   "Carrier_42_G120DControlWord.4" AT %I2460.4 : Bool;   // Bit_04_EN_RAMP
   "Carrier_42_G120DControlWord.5" AT %I2460.5 : Bool;   // Bit_05_START_RAMP
   "Carrier_42_G120DControlWord.6" AT %I2460.6 : Bool;   // Bit_06_SETPOINT
   "Carrier_42_G120DControlWord.7" AT %I2460.7 : Bool;   // Bit_07_RESET
   "Carrier_42_G120DControlWord.8" AT %I2461.0 : Bool;   // Bit_08_JOG_R
   "Carrier_42_G120DControlWord.9" AT %I2461.1 : Bool;   // Bit_09_JOG_L
   "Carrier_42_G120DControlWord.10" AT %I2461.2 : Bool;   // Bit_10_CONTR_PLC
   "Carrier_42_G120DControlWord.11" AT %I2461.3 : Bool;   // Bit_11_REVERSE
   "Carrier_42_G120DControlWord.12" AT %I2461.4 : Bool;   // Bit_12_BRAKE_RELEASE
   "Carrier_42_G120DControlWord.13" AT %I2461.5 : Bool;   // Bit_13_DDS
   "Carrier_42_G120DControlWord.14" AT %I2461.6 : Bool;   // Bit_14_DO0
   "Carrier_42_G120DControlWord.15" AT %I2461.7 : Bool;   // Bit_15_DO1
   "Carrier_42_G120DStatusWord" AT %IW2462 : Word;   // G120D_ZSW1_STATUS
   "Carrier_42_G120DStatusWord.0" AT %I2462.0 : Bool;   // Bit_00_READY_RUN
   "Carrier_42_G120DStatusWord.1" AT %I2462.1 : Bool;   // Bit_01_READY_ON
   "Carrier_42_G120DStatusWord.2" AT %I2462.2 : Bool;   // Bit_02_ENABLE
   "Carrier_42_G120DStatusWord.3" AT %I2462.3 : Bool;   // Bit_03_FAULT
   "Carrier_42_G120DStatusWord.4" AT %I2462.4 : Bool;   // Bit_04_OFF2
   "Carrier_42_G120DStatusWord.5" AT %I2462.5 : Bool;   // Bit_05_OFF3
   "Carrier_42_G120DStatusWord.6" AT %I2462.6 : Bool;   // Bit_06_LOCK_OUT
   "Carrier_42_G120DStatusWord.7" AT %I2462.7 : Bool;   // Bit_07_WARN
   "Carrier_42_G120DStatusWord.8" AT %I2463.0 : Bool;   // Bit_08_NO_DEVIATION
   "Carrier_42_G120DStatusWord.9" AT %I2463.1 : Bool;   // Bit_09_CONTR_PLC
   "Carrier_42_G120DStatusWord.10" AT %I2463.2 : Bool;   // Bit_10_F_MAX
   "Carrier_42_G120DStatusWord.11" AT %I2463.3 : Bool;   // Bit_11_LIMIT_REACHED
   "Carrier_42_G120DStatusWord.12" AT %I2463.4 : Bool;   // Bit_12_BRAKE_OPEN
   "Carrier_42_G120DStatusWord.13" AT %I2463.5 : Bool;   // Bit_13_NO_OVERTEMP
   "Carrier_42_G120DStatusWord.14" AT %I2463.6 : Bool;   // Bit_14_CW_CCW
   "Carrier_42_G120DStatusWord.15" AT %I2463.7 : Bool;   // Bit_15_OVERL
   "Carrier_42_Slot2_Input" AT %IW2464 : Word;   // SLOT 2 INPUT WORD
   "Carrier_42_CrashDetectSW" AT %I2464.0 : Bool;   // CRASH DETECT SW
   "Carrier_42_SpareSafetyInput(2_1)" AT %I2464.1 : Bool;   // SPARE SAFETY INPUT
   "Carrier_42_SpareSafetyInput(2_2)" AT %I2464.2 : Bool;   // SPARE SAFETY INPUT
   "Carrier_42_SpareSafetyInput(2_3)" AT %I2464.3 : Bool;   // SPARE SAFETY INPUT
   "Carrier_42_SpareSafetyInput(2_4)" AT %I2464.4 : Bool;   // SPARE SAFETY INPUT
   "Carrier_42_SpareSafetyInput(2_5)" AT %I2464.5 : Bool;   // SPARE SAFETY INPUT
   "Carrier_42_SpareSafetyInput(2_6)" AT %I2464.6 : Bool;   // SPARE SAFETY INPUT
   "Carrier_42_SpareSafetyInput(2_7)" AT %I2464.7 : Bool;   // SPARE SAFETY INPUT
   "Carrier_42_Slot3_SafetyOutput" AT %IW2465 : Word;   // SLOT 3 SAFETY OUTPUT WORD
   "Carrier_42_Crash_Detect_OK" AT %I2465.0 : Bool;   // CARRIER CRASH DETECT
   "Carrier_42_SpareSafetyOutput(3_1)" AT %I2465.1 : Bool;   // SPARE SAFETY OUTPUT
   "Carrier_42_SpareSafetyOutput(3_2)" AT %I2465.2 : Bool;   // SPARE SAFETY OUTPUT
   "Carrier_42_SpareSafetyOutput(3_3)" AT %I2465.3 : Bool;   // SPARE SAFETY OUTPUT
   "Carrier_42_SpareSafetyOutput(3_4)" AT %I2465.4 : Bool;   // SPARE SAFETY OUTPUT
   "Carrier_42_SpareSafetyOutput(3_5)" AT %I2465.5 : Bool;   // SPARE SAFETY OUTPUT
   "Carrier_42_SpareSafetyOutput(3_6)" AT %I2465.6 : Bool;   // SPARE SAFETY OUTPUT
   "Carrier_42_SpareSafetyOutput(3_7)" AT %I2465.7 : Bool;   // SPARE SAFETY OUTPUT
   "Carrier_42_Slot4_Input" AT %IW2466 : Word;   // SLOT 4 INPUT WORD
   "Carrier_42_480VPowerOn_MDCB1" AT %I2466.0 : Bool;   // 480 VAC POWER ON MDCB 1
   "Carrier_42_SpareInput(4_1)" AT %I2466.1 : Bool;   // SPARE INPUT
   "Carrier_42_SpareInput(4_2)" AT %I2466.2 : Bool;   // SPARE INPUT
   "Carrier_42_SitopSelectStatus" AT %I2466.3 : Bool;   // SITOP SELECT STATUS
   "Carrier_42_DCsupplyOnPSCB2" AT %I2466.4 : Bool;   // DC SUPPLY ON PSCB 2
   "Carrier_42_SpareInput(4_5)" AT %I2466.5 : Bool;   // SPARE INPUT
   "Carrier_42_SpareInput(4_6)" AT %I2466.6 : Bool;   // SPARE INPUT
   "Carrier_42_SpareInput(4_7)" AT %I2466.7 : Bool;   // SPARE INPUT
   "Carrier_42_PB1_ProdHoldLH" AT %I2467.0 : Bool;   // PB 1 PRODUCTION HOLD LH
   "Carrier_42_PB2_ResetLH" AT %I2467.1 : Bool;   // PB 2 RESET LH
   "Carrier_42_PB3_ProdHoldRH" AT %I2467.2 : Bool;   // PB 3 PRODUCTION HOLD RH
   "Carrier_42_PB4_ResetRH" AT %I2467.3 : Bool;   // PB 4 RESET RH
   "Carrier_42_SpareInput(4_14)" AT %I2467.4 : Bool;   // SPARE INPUT
   "Carrier_42_SpareInput(4_15)" AT %I2467.5 : Bool;   // SPARE INPUT
   "Carrier_42_SpareInput(4_16)" AT %I2467.6 : Bool;   // SPARE INPUT
   "Carrier_42_SpareInput(4_17)" AT %I2467.7 : Bool;   // SPARE INPUT
   "Carrier_42_Slot5_Output" AT %IW2468 : Word;   // SLOT 5 OUTPUT WORD
   "Carrier_42_IRD400_HMI_24VDC_ENABLE" AT %I2468.0 : Bool;   // IRD 400 PANEL HMI 24V DC POWER
   "Carrier_42_FaultLight_LH" AT %I2468.1 : Bool;   // FAULT LIGHT LH
   "Carrier_42_RunLight_LH" AT %I2468.2 : Bool;   // RUN LIGHT LH
   "Carrier_42_FaultLight_RH" AT %I2468.3 : Bool;   // FAULT LIGHT RH
   "Carrier_42_RunLight_RH" AT %I2468.4 : Bool;   // RUN LIGHT RH
   "Carrier_42_SpareOutput(5_5)" AT %I2468.5 : Bool;   // SPARE OUTPUT
   "Carrier_42_SpareOutput(5_6)" AT %I2468.6 : Bool;   // SPARE OUTPUT
   "Carrier_42_SpareOutput(5_7)" AT %I2468.7 : Bool;   // SPARE OUTPUT
   "Carrier_42_ActualSpeed" AT %IW2470 : Word;   // ACTUAL SPEED
   "Carrier_42_CarrierDriveAlarm" AT %IW2472 : Word;   // CARRIER DRIVE ALARM
   "Carrier_42_CarrierDriveWarning" AT %IW2474 : Word;   // CARRIER DRIVE WARNING
   "Carrier_43_Status" AT %IW2500 : Word;   // CARRIER STATUS WORD
   "Carrier_43_Status.0" AT %I2500.0 : Bool;   // HEARTBEAT
   "Carrier_43_Status.1" AT %I2500.1 : Bool;   // MANUAL
   "Carrier_43_Status.2" AT %I2500.2 : Bool;   // IN_AUTO
   "Carrier_43_Status.3" AT %I2500.3 : Bool;   // POSITIONING_COMPLETE
   "Carrier_43_Status.4" AT %I2500.4 : Bool;   // PRODUCTION HOLD
   "Carrier_43_Status.5" AT %I2500.5 : Bool;   // CARRIER MOVING FORWARD
   "Carrier_43_Status.6" AT %I2500.6 : Bool;   // CARRIER MOVING REVERSE
   "Carrier_43_Status.7" AT %I2500.7 : Bool;   // CARRIER FAULT
   "Carrier_43_Status.8" AT %I2501.0 : Bool;   // CRASH DETECT TRIPPED
   "Carrier_43_Status.9" AT %I2501.1 : Bool;
   "Carrier_43_Status.10" AT %I2501.2 : Bool;
   "Carrier_43_Status.11" AT %I2501.3 : Bool;
   "Carrier_43_Status.12" AT %I2501.4 : Bool;
   "Carrier_43_Status.13" AT %I2501.5 : Bool;
   "Carrier_43_Status.14" AT %I2501.6 : Bool;
   "Carrier_43_Status.15" AT %I2501.7 : Bool;
   "Carrier_43_SDCFaultCode" AT %IW2502 : Word;   // SDC FAULT CODE
   "Carrier_43_CarrierPosition" AT %ID2504 : DWord;   // CARRIER POSITION
   "Carrier_43_CarrierNumber" AT %IW2508 : Word;   // CARRIER NUMBER
   "Carrier_43_G120DControlWord" AT %IW2510 : Word;   // G120D_STW1_CONTROL
   "Carrier_43_G120DControlWord.0" AT %I2510.0 : Bool;   // Bit_00_ON
   "Carrier_43_G120DControlWord.1" AT %I2510.1 : Bool;   // Bit_01_AUS2_INH
   "Carrier_43_G120DControlWord.2" AT %I2510.2 : Bool;   // Bit_02_AUS3_STOP
   "Carrier_43_G120DControlWord.3" AT %I2510.3 : Bool;   // Bit_03_EN
   "Carrier_43_G120DControlWord.4" AT %I2510.4 : Bool;   // Bit_04_EN_RAMP
   "Carrier_43_G120DControlWord.5" AT %I2510.5 : Bool;   // Bit_05_START_RAMP
   "Carrier_43_G120DControlWord.6" AT %I2510.6 : Bool;   // Bit_06_SETPOINT
   "Carrier_43_G120DControlWord.7" AT %I2510.7 : Bool;   // Bit_07_RESET
   "Carrier_43_G120DControlWord.8" AT %I2511.0 : Bool;   // Bit_08_JOG_R
   "Carrier_43_G120DControlWord.9" AT %I2511.1 : Bool;   // Bit_09_JOG_L
   "Carrier_43_G120DControlWord.10" AT %I2511.2 : Bool;   // Bit_10_CONTR_PLC
   "Carrier_43_G120DControlWord.11" AT %I2511.3 : Bool;   // Bit_11_REVERSE
   "Carrier_43_G120DControlWord.12" AT %I2511.4 : Bool;   // Bit_12_BRAKE_RELEASE
   "Carrier_43_G120DControlWord.13" AT %I2511.5 : Bool;   // Bit_13_DDS
   "Carrier_43_G120DControlWord.14" AT %I2511.6 : Bool;   // Bit_14_DO0
   "Carrier_43_G120DControlWord.15" AT %I2511.7 : Bool;   // Bit_15_DO1
   "Carrier_43_G120DStatusWord" AT %IW2512 : Word;   // G120D_ZSW1_STATUS
   "Carrier_43_G120DStatusWord.0" AT %I2512.0 : Bool;   // Bit_00_READY_RUN
   "Carrier_43_G120DStatusWord.1" AT %I2512.1 : Bool;   // Bit_01_READY_ON
   "Carrier_43_G120DStatusWord.2" AT %I2512.2 : Bool;   // Bit_02_ENABLE
   "Carrier_43_G120DStatusWord.3" AT %I2512.3 : Bool;   // Bit_03_FAULT
   "Carrier_43_G120DStatusWord.4" AT %I2512.4 : Bool;   // Bit_04_OFF2
   "Carrier_43_G120DStatusWord.5" AT %I2512.5 : Bool;   // Bit_05_OFF3
   "Carrier_43_G120DStatusWord.6" AT %I2512.6 : Bool;   // Bit_06_LOCK_OUT
   "Carrier_43_G120DStatusWord.7" AT %I2512.7 : Bool;   // Bit_07_WARN
   "Carrier_43_G120DStatusWord.8" AT %I2513.0 : Bool;   // Bit_08_NO_DEVIATION
   "Carrier_43_G120DStatusWord.9" AT %I2513.1 : Bool;   // Bit_09_CONTR_PLC
   "Carrier_43_G120DStatusWord.10" AT %I2513.2 : Bool;   // Bit_10_F_MAX
   "Carrier_43_G120DStatusWord.11" AT %I2513.3 : Bool;   // Bit_11_LIMIT_REACHED
   "Carrier_43_G120DStatusWord.12" AT %I2513.4 : Bool;   // Bit_12_BRAKE_OPEN
   "Carrier_43_G120DStatusWord.13" AT %I2513.5 : Bool;   // Bit_13_NO_OVERTEMP
   "Carrier_43_G120DStatusWord.14" AT %I2513.6 : Bool;   // Bit_14_CW_CCW
   "Carrier_43_G120DStatusWord.15" AT %I2513.7 : Bool;   // Bit_15_OVERL
   "Carrier_43_Slot2_Input" AT %IW2514 : Word;   // SLOT 2 INPUT WORD
   "Carrier_43_CrashDetectSW" AT %I2514.0 : Bool;   // CRASH DETECT SW
   "Carrier_43_SpareSafetyInput(2_1)" AT %I2514.1 : Bool;   // SPARE SAFETY INPUT
   "Carrier_43_SpareSafetyInput(2_2)" AT %I2514.2 : Bool;   // SPARE SAFETY INPUT
   "Carrier_43_SpareSafetyInput(2_3)" AT %I2514.3 : Bool;   // SPARE SAFETY INPUT
   "Carrier_43_SpareSafetyInput(2_4)" AT %I2514.4 : Bool;   // SPARE SAFETY INPUT
   "Carrier_43_SpareSafetyInput(2_5)" AT %I2514.5 : Bool;   // SPARE SAFETY INPUT
   "Carrier_43_SpareSafetyInput(2_6)" AT %I2514.6 : Bool;   // SPARE SAFETY INPUT
   "Carrier_43_SpareSafetyInput(2_7)" AT %I2514.7 : Bool;   // SPARE SAFETY INPUT
   "Carrier_43_Slot3_SafetyOutput" AT %IW2515 : Word;   // SLOT 3 SAFETY OUTPUT WORD
   "Carrier_43_Crash_Detect_OK" AT %I2515.0 : Bool;   // CARRIER CRASH DETECT
   "Carrier_43_SpareSafetyOutput(3_1)" AT %I2515.1 : Bool;   // SPARE SAFETY OUTPUT
   "Carrier_43_SpareSafetyOutput(3_2)" AT %I2515.2 : Bool;   // SPARE SAFETY OUTPUT
   "Carrier_43_SpareSafetyOutput(3_3)" AT %I2515.3 : Bool;   // SPARE SAFETY OUTPUT
   "Carrier_43_SpareSafetyOutput(3_4)" AT %I2515.4 : Bool;   // SPARE SAFETY OUTPUT
   "Carrier_43_SpareSafetyOutput(3_5)" AT %I2515.5 : Bool;   // SPARE SAFETY OUTPUT
   "Carrier_43_SpareSafetyOutput(3_6)" AT %I2515.6 : Bool;   // SPARE SAFETY OUTPUT
   "Carrier_43_SpareSafetyOutput(3_7)" AT %I2515.7 : Bool;   // SPARE SAFETY OUTPUT
   "Carrier_43_Slot4_Input" AT %IW2516 : Word;   // SLOT 4 INPUT WORD
   "Carrier_43_480VPowerOn_MDCB1" AT %I2516.0 : Bool;   // 480 VAC POWER ON MDCB 1
   "Carrier_43_SpareInput(4_1)" AT %I2516.1 : Bool;   // SPARE INPUT
   "Carrier_43_SpareInput(4_2)" AT %I2516.2 : Bool;   // SPARE INPUT
   "Carrier_43_SitopSelectStatus" AT %I2516.3 : Bool;   // SITOP SELECT STATUS
   "Carrier_43_DCsupplyOnPSCB2" AT %I2516.4 : Bool;   // DC SUPPLY ON PSCB 2
   "Carrier_43_SpareInput(4_5)" AT %I2516.5 : Bool;   // SPARE INPUT
   "Carrier_43_SpareInput(4_6)" AT %I2516.6 : Bool;   // SPARE INPUT
   "Carrier_43_SpareInput(4_7)" AT %I2516.7 : Bool;   // SPARE INPUT
   "Carrier_43_PB1_ProdHoldLH" AT %I2517.0 : Bool;   // PB 1 PRODUCTION HOLD LH
   "Carrier_43_PB2_ResetLH" AT %I2517.1 : Bool;   // PB 2 RESET LH
   "Carrier_43_PB3_ProdHoldRH" AT %I2517.2 : Bool;   // PB 3 PRODUCTION HOLD RH
   "Carrier_43_PB4_ResetRH" AT %I2517.3 : Bool;   // PB 4 RESET RH
   "Carrier_43_SpareInput(4_14)" AT %I2517.4 : Bool;   // SPARE INPUT
   "Carrier_43_SpareInput(4_15)" AT %I2517.5 : Bool;   // SPARE INPUT
   "Carrier_43_SpareInput(4_16)" AT %I2517.6 : Bool;   // SPARE INPUT
   "Carrier_43_SpareInput(4_17)" AT %I2517.7 : Bool;   // SPARE INPUT
   "Carrier_43_Slot5_Output" AT %IW2518 : Word;   // SLOT 5 OUTPUT WORD
   "Carrier_43_IRD400_HMI_24VDC_ENABLE" AT %I2518.0 : Bool;   // IRD 400 PANEL HMI 24V DC POWER
   "Carrier_43_FaultLight_LH" AT %I2518.1 : Bool;   // FAULT LIGHT LH
   "Carrier_43_RunLight_LH" AT %I2518.2 : Bool;   // RUN LIGHT LH
   "Carrier_43_FaultLight_RH" AT %I2518.3 : Bool;   // FAULT LIGHT RH
   "Carrier_43_RunLight_RH" AT %I2518.4 : Bool;   // RUN LIGHT RH
   "Carrier_43_SpareOutput(5_5)" AT %I2518.5 : Bool;   // SPARE OUTPUT
   "Carrier_43_SpareOutput(5_6)" AT %I2518.6 : Bool;   // SPARE OUTPUT
   "Carrier_43_SpareOutput(5_7)" AT %I2518.7 : Bool;   // SPARE OUTPUT
   "Carrier_43_ActualSpeed" AT %IW2520 : Word;   // ACTUAL SPEED
   "Carrier_43_CarrierDriveAlarm" AT %IW2522 : Word;   // CARRIER DRIVE ALARM
   "Carrier_43_CarrierDriveWarning" AT %IW2524 : Word;   // CARRIER DRIVE WARNING
   "Carrier_44_Status" AT %IW2550 : Word;   // CARRIER STATUS WORD
   "Carrier_44_Status.0" AT %I2550.0 : Bool;   // HEARTBEAT
   "Carrier_44_Status.1" AT %I2550.1 : Bool;   // MANUAL
   "Carrier_44_Status.2" AT %I2550.2 : Bool;   // IN_AUTO
   "Carrier_44_Status.3" AT %I2550.3 : Bool;   // POSITIONING_COMPLETE
   "Carrier_44_Status.4" AT %I2550.4 : Bool;   // PRODUCTION HOLD
   "Carrier_44_Status.5" AT %I2550.5 : Bool;   // CARRIER MOVING FORWARD
   "Carrier_44_Status.6" AT %I2550.6 : Bool;   // CARRIER MOVING REVERSE
   "Carrier_44_Status.7" AT %I2550.7 : Bool;   // CARRIER FAULT
   "Carrier_44_Status.8" AT %I2551.0 : Bool;   // CRASH DETECT TRIPPED
   "Carrier_44_Status.9" AT %I2551.1 : Bool;
   "Carrier_44_Status.10" AT %I2551.2 : Bool;
   "Carrier_44_Status.11" AT %I2551.3 : Bool;
   "Carrier_44_Status.12" AT %I2551.4 : Bool;
   "Carrier_44_Status.13" AT %I2551.5 : Bool;
   "Carrier_44_Status.14" AT %I2551.6 : Bool;
   "Carrier_44_Status.15" AT %I2551.7 : Bool;
   "Carrier_44_SDCFaultCode" AT %IW2552 : Word;   // SDC FAULT CODE
   "Carrier_44_CarrierPosition" AT %ID2554 : DWord;   // CARRIER POSITION
   "Carrier_44_CarrierNumber" AT %IW2558 : Word;   // CARRIER NUMBER
   "Carrier_44_G120DControlWord" AT %IW2560 : Word;   // G120D_STW1_CONTROL
   "Carrier_44_G120DControlWord.0" AT %I2560.0 : Bool;   // Bit_00_ON
   "Carrier_44_G120DControlWord.1" AT %I2560.1 : Bool;   // Bit_01_AUS2_INH
   "Carrier_44_G120DControlWord.2" AT %I2560.2 : Bool;   // Bit_02_AUS3_STOP
   "Carrier_44_G120DControlWord.3" AT %I2560.3 : Bool;   // Bit_03_EN
   "Carrier_44_G120DControlWord.4" AT %I2560.4 : Bool;   // Bit_04_EN_RAMP
   "Carrier_44_G120DControlWord.5" AT %I2560.5 : Bool;   // Bit_05_START_RAMP
   "Carrier_44_G120DControlWord.6" AT %I2560.6 : Bool;   // Bit_06_SETPOINT
   "Carrier_44_G120DControlWord.7" AT %I2560.7 : Bool;   // Bit_07_RESET
   "Carrier_44_G120DControlWord.8" AT %I2561.0 : Bool;   // Bit_08_JOG_R
   "Carrier_44_G120DControlWord.9" AT %I2561.1 : Bool;   // Bit_09_JOG_L
   "Carrier_44_G120DControlWord.10" AT %I2561.2 : Bool;   // Bit_10_CONTR_PLC
   "Carrier_44_G120DControlWord.11" AT %I2561.3 : Bool;   // Bit_11_REVERSE
   "Carrier_44_G120DControlWord.12" AT %I2561.4 : Bool;   // Bit_12_BRAKE_RELEASE
   "Carrier_44_G120DControlWord.13" AT %I2561.5 : Bool;   // Bit_13_DDS
   "Carrier_44_G120DControlWord.14" AT %I2561.6 : Bool;   // Bit_14_DO0
   "Carrier_44_G120DControlWord.15" AT %I2561.7 : Bool;   // Bit_15_DO1
   "Carrier_44_G120DStatusWord" AT %IW2562 : Word;   // G120D_ZSW1_STATUS
   "Carrier_44_G120DStatusWord.0" AT %I2562.0 : Bool;   // Bit_00_READY_RUN
   "Carrier_44_G120DStatusWord.1" AT %I2562.1 : Bool;   // Bit_01_READY_ON
   "Carrier_44_G120DStatusWord.2" AT %I2562.2 : Bool;   // Bit_02_ENABLE
   "Carrier_44_G120DStatusWord.3" AT %I2562.3 : Bool;   // Bit_03_FAULT
   "Carrier_44_G120DStatusWord.4" AT %I2562.4 : Bool;   // Bit_04_OFF2
   "Carrier_44_G120DStatusWord.5" AT %I2562.5 : Bool;   // Bit_05_OFF3
   "Carrier_44_G120DStatusWord.6" AT %I2562.6 : Bool;   // Bit_06_LOCK_OUT
   "Carrier_44_G120DStatusWord.7" AT %I2562.7 : Bool;   // Bit_07_WARN
   "Carrier_44_G120DStatusWord.8" AT %I2563.0 : Bool;   // Bit_08_NO_DEVIATION
   "Carrier_44_G120DStatusWord.9" AT %I2563.1 : Bool;   // Bit_09_CONTR_PLC
   "Carrier_44_G120DStatusWord.10" AT %I2563.2 : Bool;   // Bit_10_F_MAX
   "Carrier_44_G120DStatusWord.11" AT %I2563.3 : Bool;   // Bit_11_LIMIT_REACHED
   "Carrier_44_G120DStatusWord.12" AT %I2563.4 : Bool;   // Bit_12_BRAKE_OPEN
   "Carrier_44_G120DStatusWord.13" AT %I2563.5 : Bool;   // Bit_13_NO_OVERTEMP
   "Carrier_44_G120DStatusWord.14" AT %I2563.6 : Bool;   // Bit_14_CW_CCW
   "Carrier_44_G120DStatusWord.15" AT %I2563.7 : Bool;   // Bit_15_OVERL
   "Carrier_44_Slot2_Input" AT %IW2564 : Word;   // SLOT 2 INPUT WORD
   "Carrier_44_CrashDetectSW" AT %I2564.0 : Bool;   // CRASH DETECT SW
   "Carrier_44_SpareSafetyInput(2_1)" AT %I2564.1 : Bool;   // SPARE SAFETY INPUT
   "Carrier_44_SpareSafetyInput(2_2)" AT %I2564.2 : Bool;   // SPARE SAFETY INPUT
   "Carrier_44_SpareSafetyInput(2_3)" AT %I2564.3 : Bool;   // SPARE SAFETY INPUT
   "Carrier_44_SpareSafetyInput(2_4)" AT %I2564.4 : Bool;   // SPARE SAFETY INPUT
   "Carrier_44_SpareSafetyInput(2_5)" AT %I2564.5 : Bool;   // SPARE SAFETY INPUT
   "Carrier_44_SpareSafetyInput(2_6)" AT %I2564.6 : Bool;   // SPARE SAFETY INPUT
   "Carrier_44_SpareSafetyInput(2_7)" AT %I2564.7 : Bool;   // SPARE SAFETY INPUT
   "Carrier_44_Slot3_SafetyOutput" AT %IW2565 : Word;   // SLOT 3 SAFETY OUTPUT WORD
   "Carrier_44_Crash_Detect_OK" AT %I2565.0 : Bool;   // CARRIER CRASH DETECT
   "Carrier_44_SpareSafetyOutput(3_1)" AT %I2565.1 : Bool;   // SPARE SAFETY OUTPUT
   "Carrier_44_SpareSafetyOutput(3_2)" AT %I2565.2 : Bool;   // SPARE SAFETY OUTPUT
   "Carrier_44_SpareSafetyOutput(3_3)" AT %I2565.3 : Bool;   // SPARE SAFETY OUTPUT
   "Carrier_44_SpareSafetyOutput(3_4)" AT %I2565.4 : Bool;   // SPARE SAFETY OUTPUT
   "Carrier_44_SpareSafetyOutput(3_5)" AT %I2565.5 : Bool;   // SPARE SAFETY OUTPUT
   "Carrier_44_SpareSafetyOutput(3_6)" AT %I2565.6 : Bool;   // SPARE SAFETY OUTPUT
   "Carrier_44_SpareSafetyOutput(3_7)" AT %I2565.7 : Bool;   // SPARE SAFETY OUTPUT
   "Carrier_44_Slot4_Input" AT %IW2566 : Word;   // SLOT 4 INPUT WORD
   "Carrier_44_480VPowerOn_MDCB1" AT %I2566.0 : Bool;   // 480 VAC POWER ON MDCB 1
   "Carrier_44_SpareInput(4_1)" AT %I2566.1 : Bool;   // SPARE INPUT
   "Carrier_44_SpareInput(4_2)" AT %I2566.2 : Bool;   // SPARE INPUT
   "Carrier_44_SitopSelectStatus" AT %I2566.3 : Bool;   // SITOP SELECT STATUS
   "Carrier_44_DCsupplyOnPSCB2" AT %I2566.4 : Bool;   // DC SUPPLY ON PSCB 2
   "Carrier_44_SpareInput(4_5)" AT %I2566.5 : Bool;   // SPARE INPUT
   "Carrier_44_SpareInput(4_6)" AT %I2566.6 : Bool;   // SPARE INPUT
   "Carrier_44_SpareInput(4_7)" AT %I2566.7 : Bool;   // SPARE INPUT
   "Carrier_44_PB1_ProdHoldLH" AT %I2567.0 : Bool;   // PB 1 PRODUCTION HOLD LH
   "Carrier_44_PB2_ResetLH" AT %I2567.1 : Bool;   // PB 2 RESET LH
   "Carrier_44_PB3_ProdHoldRH" AT %I2567.2 : Bool;   // PB 3 PRODUCTION HOLD RH
   "Carrier_44_PB4_ResetRH" AT %I2567.3 : Bool;   // PB 4 RESET RH
   "Carrier_44_SpareInput(4_14)" AT %I2567.4 : Bool;   // SPARE INPUT
   "Carrier_44_SpareInput(4_15)" AT %I2567.5 : Bool;   // SPARE INPUT
   "Carrier_44_SpareInput(4_16)" AT %I2567.6 : Bool;   // SPARE INPUT
   "Carrier_44_SpareInput(4_17)" AT %I2567.7 : Bool;   // SPARE INPUT
   "Carrier_44_Slot5_Output" AT %IW2568 : Word;   // SLOT 5 OUTPUT WORD
   "Carrier_44_IRD400_HMI_24VDC_ENABLE" AT %I2568.0 : Bool;   // IRD 400 PANEL HMI 24V DC POWER
   "Carrier_44_FaultLight_LH" AT %I2568.1 : Bool;   // FAULT LIGHT LH
   "Carrier_44_RunLight_LH" AT %I2568.2 : Bool;   // RUN LIGHT LH
   "Carrier_44_FaultLight_RH" AT %I2568.3 : Bool;   // FAULT LIGHT RH
   "Carrier_44_RunLight_RH" AT %I2568.4 : Bool;   // RUN LIGHT RH
   "Carrier_44_SpareOutput(5_5)" AT %I2568.5 : Bool;   // SPARE OUTPUT
   "Carrier_44_SpareOutput(5_6)" AT %I2568.6 : Bool;   // SPARE OUTPUT
   "Carrier_44_SpareOutput(5_7)" AT %I2568.7 : Bool;   // SPARE OUTPUT
   "Carrier_44_ActualSpeed" AT %IW2570 : Word;   // ACTUAL SPEED
   "Carrier_44_CarrierDriveAlarm" AT %IW2572 : Word;   // CARRIER DRIVE ALARM
   "Carrier_44_CarrierDriveWarning" AT %IW2574 : Word;   // CARRIER DRIVE WARNING
   "Carrier_45_Status" AT %IW2600 : Word;   // CARRIER STATUS WORD
   "Carrier_45_Status.0" AT %I2600.0 : Bool;   // HEARTBEAT
   "Carrier_45_Status.1" AT %I2600.1 : Bool;   // MANUAL
   "Carrier_45_Status.2" AT %I2600.2 : Bool;   // IN_AUTO
   "Carrier_45_Status.3" AT %I2600.3 : Bool;   // POSITIONING_COMPLETE
   "Carrier_45_Status.4" AT %I2600.4 : Bool;   // PRODUCTION HOLD
   "Carrier_45_Status.5" AT %I2600.5 : Bool;   // CARRIER MOVING FORWARD
   "Carrier_45_Status.6" AT %I2600.6 : Bool;   // CARRIER MOVING REVERSE
   "Carrier_45_Status.7" AT %I2600.7 : Bool;   // CARRIER FAULT
   "Carrier_45_Status.8" AT %I2601.0 : Bool;   // CRASH DETECT TRIPPED
   "Carrier_45_Status.9" AT %I2601.1 : Bool;
   "Carrier_45_Status.10" AT %I2601.2 : Bool;
   "Carrier_45_Status.11" AT %I2601.3 : Bool;
   "Carrier_45_Status.12" AT %I2601.4 : Bool;
   "Carrier_45_Status.13" AT %I2601.5 : Bool;
   "Carrier_45_Status.14" AT %I2601.6 : Bool;
   "Carrier_45_Status.15" AT %I2601.7 : Bool;
   "Carrier_45_SDCFaultCode" AT %IW2602 : Word;   // SDC FAULT CODE
   "Carrier_45_CarrierPosition" AT %ID2604 : DWord;   // CARRIER POSITION
   "Carrier_45_CarrierNumber" AT %IW2608 : Word;   // CARRIER NUMBER
   "Carrier_45_G120DControlWord" AT %IW2610 : Word;   // G120D_STW1_CONTROL
   "Carrier_45_G120DControlWord.0" AT %I2610.0 : Bool;   // Bit_00_ON
   "Carrier_45_G120DControlWord.1" AT %I2610.1 : Bool;   // Bit_01_AUS2_INH
   "Carrier_45_G120DControlWord.2" AT %I2610.2 : Bool;   // Bit_02_AUS3_STOP
   "Carrier_45_G120DControlWord.3" AT %I2610.3 : Bool;   // Bit_03_EN
   "Carrier_45_G120DControlWord.4" AT %I2610.4 : Bool;   // Bit_04_EN_RAMP
   "Carrier_45_G120DControlWord.5" AT %I2610.5 : Bool;   // Bit_05_START_RAMP
   "Carrier_45_G120DControlWord.6" AT %I2610.6 : Bool;   // Bit_06_SETPOINT
   "Carrier_45_G120DControlWord.7" AT %I2610.7 : Bool;   // Bit_07_RESET
   "Carrier_45_G120DControlWord.8" AT %I2611.0 : Bool;   // Bit_08_JOG_R
   "Carrier_45_G120DControlWord.9" AT %I2611.1 : Bool;   // Bit_09_JOG_L
   "Carrier_45_G120DControlWord.10" AT %I2611.2 : Bool;   // Bit_10_CONTR_PLC
   "Carrier_45_G120DControlWord.11" AT %I2611.3 : Bool;   // Bit_11_REVERSE
   "Carrier_45_G120DControlWord.12" AT %I2611.4 : Bool;   // Bit_12_BRAKE_RELEASE
   "Carrier_45_G120DControlWord.13" AT %I2611.5 : Bool;   // Bit_13_DDS
   "Carrier_45_G120DControlWord.14" AT %I2611.6 : Bool;   // Bit_14_DO0
   "Carrier_45_G120DControlWord.15" AT %I2611.7 : Bool;   // Bit_15_DO1
   "Carrier_45_G120DStatusWord" AT %IW2612 : Word;   // G120D_ZSW1_STATUS
   "Carrier_45_G120DStatusWord.0" AT %I2612.0 : Bool;   // Bit_00_READY_RUN
   "Carrier_45_G120DStatusWord.1" AT %I2612.1 : Bool;   // Bit_01_READY_ON
   "Carrier_45_G120DStatusWord.2" AT %I2612.2 : Bool;   // Bit_02_ENABLE
   "Carrier_45_G120DStatusWord.3" AT %I2612.3 : Bool;   // Bit_03_FAULT
   "Carrier_45_G120DStatusWord.4" AT %I2612.4 : Bool;   // Bit_04_OFF2
   "Carrier_45_G120DStatusWord.5" AT %I2612.5 : Bool;   // Bit_05_OFF3
   "Carrier_45_G120DStatusWord.6" AT %I2612.6 : Bool;   // Bit_06_LOCK_OUT
   "Carrier_45_G120DStatusWord.7" AT %I2612.7 : Bool;   // Bit_07_WARN
   "Carrier_45_G120DStatusWord.8" AT %I2613.0 : Bool;   // Bit_08_NO_DEVIATION
   "Carrier_45_G120DStatusWord.9" AT %I2613.1 : Bool;   // Bit_09_CONTR_PLC
   "Carrier_45_G120DStatusWord.10" AT %I2613.2 : Bool;   // Bit_10_F_MAX
   "Carrier_45_G120DStatusWord.11" AT %I2613.3 : Bool;   // Bit_11_LIMIT_REACHED
   "Carrier_45_G120DStatusWord.12" AT %I2613.4 : Bool;   // Bit_12_BRAKE_OPEN
   "Carrier_45_G120DStatusWord.13" AT %I2613.5 : Bool;   // Bit_13_NO_OVERTEMP
   "Carrier_45_G120DStatusWord.14" AT %I2613.6 : Bool;   // Bit_14_CW_CCW
   "Carrier_45_G120DStatusWord.15" AT %I2613.7 : Bool;   // Bit_15_OVERL
   "Carrier_45_Slot2_Input" AT %IW2614 : Word;   // SLOT 2 INPUT WORD
   "Carrier_45_CrashDetectSW" AT %I2614.0 : Bool;   // CRASH DETECT SW
   "Carrier_45_SpareSafetyInput(2_1)" AT %I2614.1 : Bool;   // SPARE SAFETY INPUT
   "Carrier_45_SpareSafetyInput(2_2)" AT %I2614.2 : Bool;   // SPARE SAFETY INPUT
   "Carrier_45_SpareSafetyInput(2_3)" AT %I2614.3 : Bool;   // SPARE SAFETY INPUT
   "Carrier_45_SpareSafetyInput(2_4)" AT %I2614.4 : Bool;   // SPARE SAFETY INPUT
   "Carrier_45_SpareSafetyInput(2_5)" AT %I2614.5 : Bool;   // SPARE SAFETY INPUT
   "Carrier_45_SpareSafetyInput(2_6)" AT %I2614.6 : Bool;   // SPARE SAFETY INPUT
   "Carrier_45_SpareSafetyInput(2_7)" AT %I2614.7 : Bool;   // SPARE SAFETY INPUT
   "Carrier_45_Slot3_SafetyOutput" AT %IW2615 : Word;   // SLOT 3 SAFETY OUTPUT WORD
   "Carrier_45_Crash_Detect_OK" AT %I2615.0 : Bool;   // CARRIER CRASH DETECT
   "Carrier_45_SpareSafetyOutput(3_1)" AT %I2615.1 : Bool;   // SPARE SAFETY OUTPUT
   "Carrier_45_SpareSafetyOutput(3_2)" AT %I2615.2 : Bool;   // SPARE SAFETY OUTPUT
   "Carrier_45_SpareSafetyOutput(3_3)" AT %I2615.3 : Bool;   // SPARE SAFETY OUTPUT
   "Carrier_45_SpareSafetyOutput(3_4)" AT %I2615.4 : Bool;   // SPARE SAFETY OUTPUT
   "Carrier_45_SpareSafetyOutput(3_5)" AT %I2615.5 : Bool;   // SPARE SAFETY OUTPUT
   "Carrier_45_SpareSafetyOutput(3_6)" AT %I2615.6 : Bool;   // SPARE SAFETY OUTPUT
   "Carrier_45_SpareSafetyOutput(3_7)" AT %I2615.7 : Bool;   // SPARE SAFETY OUTPUT
   "Carrier_45_Slot4_Input" AT %IW2616 : Word;   // SLOT 4 INPUT WORD
   "Carrier_45_480VPowerOn_MDCB1" AT %I2616.0 : Bool;   // 480 VAC POWER ON MDCB 1
   "Carrier_45_SpareInput(4_1)" AT %I2616.1 : Bool;   // SPARE INPUT
   "Carrier_45_SpareInput(4_2)" AT %I2616.2 : Bool;   // SPARE INPUT
   "Carrier_45_SitopSelectStatus" AT %I2616.3 : Bool;   // SITOP SELECT STATUS
   "Carrier_45_DCsupplyOnPSCB2" AT %I2616.4 : Bool;   // DC SUPPLY ON PSCB 2
   "Carrier_45_SpareInput(4_5)" AT %I2616.5 : Bool;   // SPARE INPUT
   "Carrier_45_SpareInput(4_6)" AT %I2616.6 : Bool;   // SPARE INPUT
   "Carrier_45_SpareInput(4_7)" AT %I2616.7 : Bool;   // SPARE INPUT
   "Carrier_45_PB1_ProdHoldLH" AT %I2617.0 : Bool;   // PB 1 PRODUCTION HOLD LH
   "Carrier_45_PB2_ResetLH" AT %I2617.1 : Bool;   // PB 2 RESET LH
   "Carrier_45_PB3_ProdHoldRH" AT %I2617.2 : Bool;   // PB 3 PRODUCTION HOLD RH
   "Carrier_45_PB4_ResetRH" AT %I2617.3 : Bool;   // PB 4 RESET RH
   "Carrier_45_SpareInput(4_14)" AT %I2617.4 : Bool;   // SPARE INPUT
   "Carrier_45_SpareInput(4_15)" AT %I2617.5 : Bool;   // SPARE INPUT
   "Carrier_45_SpareInput(4_16)" AT %I2617.6 : Bool;   // SPARE INPUT
   "Carrier_45_SpareInput(4_17)" AT %I2617.7 : Bool;   // SPARE INPUT
   "Carrier_45_Slot5_Output" AT %IW2618 : Word;   // SLOT 5 OUTPUT WORD
   "Carrier_45_IRD400_HMI_24VDC_ENABLE" AT %I2618.0 : Bool;   // IRD 400 PANEL HMI 24V DC POWER
   "Carrier_45_FaultLight_LH" AT %I2618.1 : Bool;   // FAULT LIGHT LH
   "Carrier_45_RunLight_LH" AT %I2618.2 : Bool;   // RUN LIGHT LH
   "Carrier_45_FaultLight_RH" AT %I2618.3 : Bool;   // FAULT LIGHT RH
   "Carrier_45_RunLight_RH" AT %I2618.4 : Bool;   // RUN LIGHT RH
   "Carrier_45_SpareOutput(5_5)" AT %I2618.5 : Bool;   // SPARE OUTPUT
   "Carrier_45_SpareOutput(5_6)" AT %I2618.6 : Bool;   // SPARE OUTPUT
   "Carrier_45_SpareOutput(5_7)" AT %I2618.7 : Bool;   // SPARE OUTPUT
   "Carrier_45_ActualSpeed" AT %IW2620 : Word;   // ACTUAL SPEED
   "Carrier_45_CarrierDriveAlarm" AT %IW2622 : Word;   // CARRIER DRIVE ALARM
   "Carrier_45_CarrierDriveWarning" AT %IW2624 : Word;   // CARRIER DRIVE WARNING
   "Carrier_46_Status" AT %IW2650 : Word;   // CARRIER STATUS WORD
   "Carrier_46_Status.0" AT %I2650.0 : Bool;   // HEARTBEAT
   "Carrier_46_Status.1" AT %I2650.1 : Bool;   // MANUAL
   "Carrier_46_Status.2" AT %I2650.2 : Bool;   // IN_AUTO
   "Carrier_46_Status.3" AT %I2650.3 : Bool;   // POSITIONING_COMPLETE
   "Carrier_46_Status.4" AT %I2650.4 : Bool;   // PRODUCTION HOLD
   "Carrier_46_Status.5" AT %I2650.5 : Bool;   // CARRIER MOVING FORWARD
   "Carrier_46_Status.6" AT %I2650.6 : Bool;   // CARRIER MOVING REVERSE
   "Carrier_46_Status.7" AT %I2650.7 : Bool;   // CARRIER FAULT
   "Carrier_46_Status.8" AT %I2651.0 : Bool;   // CRASH DETECT TRIPPED
   "Carrier_46_Status.9" AT %I2651.1 : Bool;
   "Carrier_46_Status.10" AT %I2651.2 : Bool;
   "Carrier_46_Status.11" AT %I2651.3 : Bool;
   "Carrier_46_Status.12" AT %I2651.4 : Bool;
   "Carrier_46_Status.13" AT %I2651.5 : Bool;
   "Carrier_46_Status.14" AT %I2651.6 : Bool;
   "Carrier_46_Status.15" AT %I2651.7 : Bool;
   "Carrier_46_SDCFaultCode" AT %IW2652 : Word;   // SDC FAULT CODE
   "Carrier_46_CarrierPosition" AT %ID2654 : DWord;   // CARRIER POSITION
   "Carrier_46_CarrierNumber" AT %IW2658 : Word;   // CARRIER NUMBER
   "Carrier_46_G120DControlWord" AT %IW2660 : Word;   // G120D_STW1_CONTROL
   "Carrier_46_G120DControlWord.0" AT %I2660.0 : Bool;   // Bit_00_ON
   "Carrier_46_G120DControlWord.1" AT %I2660.1 : Bool;   // Bit_01_AUS2_INH
   "Carrier_46_G120DControlWord.2" AT %I2660.2 : Bool;   // Bit_02_AUS3_STOP
   "Carrier_46_G120DControlWord.3" AT %I2660.3 : Bool;   // Bit_03_EN
   "Carrier_46_G120DControlWord.4" AT %I2660.4 : Bool;   // Bit_04_EN_RAMP
   "Carrier_46_G120DControlWord.5" AT %I2660.5 : Bool;   // Bit_05_START_RAMP
   "Carrier_46_G120DControlWord.6" AT %I2660.6 : Bool;   // Bit_06_SETPOINT
   "Carrier_46_G120DControlWord.7" AT %I2660.7 : Bool;   // Bit_07_RESET
   "Carrier_46_G120DControlWord.8" AT %I2661.0 : Bool;   // Bit_08_JOG_R
   "Carrier_46_G120DControlWord.9" AT %I2661.1 : Bool;   // Bit_09_JOG_L
   "Carrier_46_G120DControlWord.10" AT %I2661.2 : Bool;   // Bit_10_CONTR_PLC
   "Carrier_46_G120DControlWord.11" AT %I2661.3 : Bool;   // Bit_11_REVERSE
   "Carrier_46_G120DControlWord.12" AT %I2661.4 : Bool;   // Bit_12_BRAKE_RELEASE
   "Carrier_46_G120DControlWord.13" AT %I2661.5 : Bool;   // Bit_13_DDS
   "Carrier_46_G120DControlWord.14" AT %I2661.6 : Bool;   // Bit_14_DO0
   "Carrier_46_G120DControlWord.15" AT %I2661.7 : Bool;   // Bit_15_DO1
   "Carrier_46_G120DStatusWord" AT %IW2662 : Word;   // G120D_ZSW1_STATUS
   "Carrier_46_G120DStatusWord.0" AT %I2662.0 : Bool;   // Bit_00_READY_RUN
   "Carrier_46_G120DStatusWord.1" AT %I2662.1 : Bool;   // Bit_01_READY_ON
   "Carrier_46_G120DStatusWord.2" AT %I2662.2 : Bool;   // Bit_02_ENABLE
   "Carrier_46_G120DStatusWord.3" AT %I2662.3 : Bool;   // Bit_03_FAULT
   "Carrier_46_G120DStatusWord.4" AT %I2662.4 : Bool;   // Bit_04_OFF2
   "Carrier_46_G120DStatusWord.5" AT %I2662.5 : Bool;   // Bit_05_OFF3
   "Carrier_46_G120DStatusWord.6" AT %I2662.6 : Bool;   // Bit_06_LOCK_OUT
   "Carrier_46_G120DStatusWord.7" AT %I2662.7 : Bool;   // Bit_07_WARN
   "Carrier_46_G120DStatusWord.8" AT %I2663.0 : Bool;   // Bit_08_NO_DEVIATION
   "Carrier_46_G120DStatusWord.9" AT %I2663.1 : Bool;   // Bit_09_CONTR_PLC
   "Carrier_46_G120DStatusWord.10" AT %I2663.2 : Bool;   // Bit_10_F_MAX
   "Carrier_46_G120DStatusWord.11" AT %I2663.3 : Bool;   // Bit_11_LIMIT_REACHED
   "Carrier_46_G120DStatusWord.12" AT %I2663.4 : Bool;   // Bit_12_BRAKE_OPEN
   "Carrier_46_G120DStatusWord.13" AT %I2663.5 : Bool;   // Bit_13_NO_OVERTEMP
   "Carrier_46_G120DStatusWord.14" AT %I2663.6 : Bool;   // Bit_14_CW_CCW
   "Carrier_46_G120DStatusWord.15" AT %I2663.7 : Bool;   // Bit_15_OVERL
   "Carrier_46_Slot2_Input" AT %IW2664 : Word;   // SLOT 2 INPUT WORD
   "Carrier_46_CrashDetectSW" AT %I2664.0 : Bool;   // CRASH DETECT SW
   "Carrier_46_SpareSafetyInput(2_1)" AT %I2664.1 : Bool;   // SPARE SAFETY INPUT
   "Carrier_46_SpareSafetyInput(2_2)" AT %I2664.2 : Bool;   // SPARE SAFETY INPUT
   "Carrier_46_SpareSafetyInput(2_3)" AT %I2664.3 : Bool;   // SPARE SAFETY INPUT
   "Carrier_46_SpareSafetyInput(2_4)" AT %I2664.4 : Bool;   // SPARE SAFETY INPUT
   "Carrier_46_SpareSafetyInput(2_5)" AT %I2664.5 : Bool;   // SPARE SAFETY INPUT
   "Carrier_46_SpareSafetyInput(2_6)" AT %I2664.6 : Bool;   // SPARE SAFETY INPUT
   "Carrier_46_SpareSafetyInput(2_7)" AT %I2664.7 : Bool;   // SPARE SAFETY INPUT
   "Carrier_46_Slot3_SafetyOutput" AT %IW2665 : Word;   // SLOT 3 SAFETY OUTPUT WORD
   "Carrier_46_Crash_Detect_OK" AT %I2665.0 : Bool;   // CARRIER CRASH DETECT
   "Carrier_46_SpareSafetyOutput(3_1)" AT %I2665.1 : Bool;   // SPARE SAFETY OUTPUT
   "Carrier_46_SpareSafetyOutput(3_2)" AT %I2665.2 : Bool;   // SPARE SAFETY OUTPUT
   "Carrier_46_SpareSafetyOutput(3_3)" AT %I2665.3 : Bool;   // SPARE SAFETY OUTPUT
   "Carrier_46_SpareSafetyOutput(3_4)" AT %I2665.4 : Bool;   // SPARE SAFETY OUTPUT
   "Carrier_46_SpareSafetyOutput(3_5)" AT %I2665.5 : Bool;   // SPARE SAFETY OUTPUT
   "Carrier_46_SpareSafetyOutput(3_6)" AT %I2665.6 : Bool;   // SPARE SAFETY OUTPUT
   "Carrier_46_SpareSafetyOutput(3_7)" AT %I2665.7 : Bool;   // SPARE SAFETY OUTPUT
   "Carrier_46_Slot4_Input" AT %IW2666 : Word;   // SLOT 4 INPUT WORD
   "Carrier_46_480VPowerOn_MDCB1" AT %I2666.0 : Bool;   // 480 VAC POWER ON MDCB 1
   "Carrier_46_SpareInput(4_1)" AT %I2666.1 : Bool;   // SPARE INPUT
   "Carrier_46_SpareInput(4_2)" AT %I2666.2 : Bool;   // SPARE INPUT
   "Carrier_46_SitopSelectStatus" AT %I2666.3 : Bool;   // SITOP SELECT STATUS
   "Carrier_46_DCsupplyOnPSCB2" AT %I2666.4 : Bool;   // DC SUPPLY ON PSCB 2
   "Carrier_46_SpareInput(4_5)" AT %I2666.5 : Bool;   // SPARE INPUT